VERSION : 0.1
   VAR
      HEADER : Struct
         DB_NR : Int := 3701;
         MIN_NR_EMS : Int := 1;
         MAX_NR_EMS : Int := 200;
         START_EMS : Int := 20;
         LAENGE_EMS_FLAGS : Int := 2;
         ACT_COUNT : Int := 0;
         Res120 : Int := 0;
         Res140 : Int := 0;
         Res160 : Int := 0;
         Res180 : Int := 0;
      END_STRUCT;
      EMS : Array[1..200] of "UDT_SDC_EMS_FLAGS";
      LADDR_EMS : Array[1..200] of HW_ANY;
   END_VAR
BEGIN
   EMS[3].SIMULATION := FALSE;
   EMS[2].SIMULATION := FALSE;
   EMS[200].FAULTY := TRUE;
   EMS[199].FAULTY := TRUE;
   EMS[198].FAULTY := TRUE;
   EMS[197].FAULTY := TRUE;
   EMS[196].FAULTY := TRUE;
   EMS[195].FAULTY := TRUE;
   EMS[194].FAULTY := TRUE;
   EMS[193].FAULTY := TRUE;
   EMS[192].FAULTY := TRUE;
   EMS[191].FAULTY := TRUE;
   EMS[190].FAULTY := TRUE;
   EMS[189].FAULTY := TRUE;
   EMS[188].FAULTY := TRUE;
   EMS[187].FAULTY := TRUE;
   EMS[186].FAULTY := TRUE;
   EMS[185].FAULTY := TRUE;
   EMS[184].FAULTY := TRUE;
   EMS[183].FAULTY := TRUE;
   EMS[182].FAULTY := TRUE;
   EMS[181].FAULTY := TRUE;
   EMS[180].FAULTY := TRUE;
   EMS[179].FAULTY := TRUE;
   EMS[178].FAULTY := TRUE;
   EMS[177].FAULTY := TRUE;
   EMS[176].FAULTY := TRUE;
   EMS[175].FAULTY := TRUE;
   EMS[174].FAULTY := TRUE;
   EMS[173].FAULTY := TRUE;
   EMS[172].FAULTY := TRUE;
   EMS[171].FAULTY := TRUE;
   EMS[170].FAULTY := TRUE;
   EMS[169].FAULTY := TRUE;
   EMS[168].FAULTY := TRUE;
   EMS[167].FAULTY := TRUE;
   EMS[166].FAULTY := TRUE;
   EMS[165].FAULTY := TRUE;
   EMS[164].FAULTY := TRUE;
   EMS[163].FAULTY := TRUE;
   EMS[162].FAULTY := TRUE;
   EMS[161].FAULTY := TRUE;
   EMS[160].FAULTY := TRUE;
   EMS[159].FAULTY := TRUE;
   EMS[158].FAULTY := TRUE;
   EMS[157].FAULTY := TRUE;
   EMS[156].FAULTY := TRUE;
   EMS[155].FAULTY := TRUE;
   EMS[154].FAULTY := TRUE;
   EMS[153].FAULTY := TRUE;
   EMS[152].FAULTY := TRUE;
   EMS[151].FAULTY := TRUE;
   EMS[150].FAULTY := TRUE;
   EMS[149].FAULTY := TRUE;
   EMS[148].FAULTY := TRUE;
   EMS[147].FAULTY := TRUE;
   EMS[146].FAULTY := TRUE;
   EMS[145].FAULTY := TRUE;
   EMS[144].FAULTY := TRUE;
   EMS[143].FAULTY := TRUE;
   EMS[142].FAULTY := TRUE;
   EMS[141].FAULTY := TRUE;
   EMS[140].FAULTY := TRUE;
   EMS[139].FAULTY := TRUE;
   EMS[138].FAULTY := TRUE;
   EMS[137].FAULTY := TRUE;
   EMS[136].FAULTY := TRUE;
   EMS[135].FAULTY := TRUE;
   EMS[134].FAULTY := TRUE;
   EMS[133].FAULTY := TRUE;
   EMS[132].FAULTY := TRUE;
   EMS[131].FAULTY := TRUE;
   EMS[130].FAULTY := TRUE;
   EMS[129].FAULTY := TRUE;
   EMS[128].FAULTY := TRUE;
   EMS[127].FAULTY := TRUE;
   EMS[126].FAULTY := TRUE;
   EMS[125].FAULTY := TRUE;
   EMS[124].FAULTY := TRUE;
   EMS[123].FAULTY := TRUE;
   EMS[122].FAULTY := TRUE;
   EMS[121].FAULTY := TRUE;
   EMS[120].FAULTY := TRUE;
   EMS[119].FAULTY := TRUE;
   EMS[118].FAULTY := TRUE;
   EMS[117].FAULTY := TRUE;
   EMS[116].FAULTY := TRUE;
   EMS[115].FAULTY := TRUE;
   EMS[114].FAULTY := TRUE;
   EMS[113].FAULTY := TRUE;
   EMS[112].FAULTY := TRUE;
   EMS[111].FAULTY := TRUE;
   EMS[110].FAULTY := TRUE;
   EMS[109].FAULTY := TRUE;
   EMS[108].FAULTY := TRUE;
   EMS[107].FAULTY := TRUE;
   EMS[106].FAULTY := TRUE;
   EMS[105].FAULTY := TRUE;
   EMS[104].FAULTY := TRUE;
   EMS[103].FAULTY := TRUE;
   EMS[102].FAULTY := TRUE;
   EMS[101].FAULTY := TRUE;
   EMS[100].FAULTY := TRUE;
   EMS[99].FAULTY := TRUE;
   EMS[98].FAULTY := TRUE;
   EMS[97].FAULTY := TRUE;
   EMS[96].FAULTY := TRUE;
   EMS[95].FAULTY := TRUE;
   EMS[94].FAULTY := TRUE;
   EMS[93].FAULTY := TRUE;
   EMS[92].FAULTY := TRUE;
   EMS[91].FAULTY := TRUE;
   EMS[90].FAULTY := TRUE;
   EMS[89].FAULTY := TRUE;
   EMS[88].FAULTY := TRUE;
   EMS[87].FAULTY := TRUE;
   EMS[86].FAULTY := TRUE;
   EMS[85].FAULTY := TRUE;
   EMS[84].FAULTY := TRUE;
   EMS[83].FAULTY := TRUE;
   EMS[82].FAULTY := TRUE;
   EMS[81].FAULTY := TRUE;
   EMS[80].FAULTY := TRUE;
   EMS[79].FAULTY := TRUE;
   EMS[78].FAULTY := TRUE;
   EMS[77].FAULTY := TRUE;
   EMS[76].FAULTY := TRUE;
   EMS[75].FAULTY := TRUE;
   EMS[74].FAULTY := TRUE;
   EMS[73].FAULTY := TRUE;
   EMS[72].FAULTY := TRUE;
   EMS[71].FAULTY := TRUE;
   EMS[70].FAULTY := TRUE;
   EMS[69].FAULTY := TRUE;
   EMS[68].FAULTY := TRUE;
   EMS[67].FAULTY := TRUE;
   EMS[66].FAULTY := TRUE;
   EMS[65].FAULTY := TRUE;
   EMS[64].FAULTY := TRUE;
   EMS[63].FAULTY := TRUE;
   EMS[62].FAULTY := TRUE;
   EMS[61].FAULTY := TRUE;
   EMS[60].FAULTY := TRUE;
   EMS[59].FAULTY := TRUE;
   EMS[58].FAULTY := TRUE;
   EMS[57].FAULTY := TRUE;
   EMS[56].FAULTY := TRUE;
   EMS[55].FAULTY := TRUE;
   EMS[54].FAULTY := FALSE;
   EMS[53].FAULTY := TRUE;
   EMS[52].FAULTY := TRUE;
   EMS[51].FAULTY := TRUE;
   EMS[50].FAULTY := TRUE;
   EMS[49].FAULTY := TRUE;
   EMS[48].FAULTY := TRUE;
   EMS[47].FAULTY := TRUE;
   EMS[46].FAULTY := TRUE;
   EMS[45].FAULTY := TRUE;
   EMS[44].FAULTY := TRUE;
   EMS[43].FAULTY := TRUE;
   EMS[42].FAULTY := TRUE;
   EMS[41].FAULTY := TRUE;
   EMS[40].FAULTY := TRUE;
   EMS[39].FAULTY := TRUE;
   EMS[38].FAULTY := TRUE;
   EMS[37].FAULTY := TRUE;
   EMS[36].FAULTY := TRUE;
   EMS[35].FAULTY := TRUE;
   EMS[34].FAULTY := FALSE;
   EMS[33].FAULTY := TRUE;
   EMS[32].FAULTY := FALSE;
   EMS[31].FAULTY := TRUE;
   EMS[30].FAULTY := TRUE;
   EMS[29].FAULTY := FALSE;
   EMS[28].FAULTY := TRUE;
   EMS[27].FAULTY := TRUE;
   EMS[26].FAULTY := TRUE;
   EMS[25].FAULTY := TRUE;
   EMS[24].FAULTY := TRUE;
   EMS[23].FAULTY := TRUE;
   EMS[22].FAULTY := TRUE;
   EMS[21].FAULTY := TRUE;
   EMS[20].FAULTY := TRUE;
   EMS[19].FAULTY := TRUE;
   EMS[18].FAULTY := TRUE;
   EMS[17].FAULTY := TRUE;
   EMS[16].FAULTY := TRUE;
   EMS[15].FAULTY := TRUE;
   EMS[14].FAULTY := TRUE;
   EMS[13].FAULTY := TRUE;
   EMS[12].FAULTY := TRUE;
   EMS[11].FAULTY := TRUE;
   EMS[10].FAULTY := TRUE;
   EMS[9].FAULTY := TRUE;
   EMS[8].FAULTY := TRUE;
   EMS[7].FAULTY := TRUE;
   EMS[6].FAULTY := TRUE;
   EMS[5].FAULTY := TRUE;
   EMS[4].FAULTY := TRUE;
   EMS[3].FAULTY := TRUE;
   // 3200 more start values not shown
END_DATA_BLOCK

DATA_BLOCK "DB_SDC_TS_PARAMETER_1"   // DB3704
{ S7_Optimized_Access := 'FALSE' }
AUTHOR : FFM
FAMILY : SDC
NAME : SECT_DEF
VERSION : 1.0
   VAR
      HEADER : Struct
         DB_NR : Int := 3704;
         MIN_NR_SEK : Int := 1;
         MAX_NR_SEK : Int := 100;
         START_DAT : Int := 20;
         LAENGE_SEK_DATA : Int := 260;
         ANZ_PROFIL : Int := 10;
         OFFEST_PROFIL : Int := 40;
         LAENGE_PROFIL_DATA : Int := 22;
         Res160 : Int := 0;
         Res : Int := 0;
      END_STRUCT;
      TS : Array[1..100] of "UDT_SDC_TS_PARAMETER";
   END_VAR
BEGIN
   TS[100].ALLG.Drive_speed_2 := 15000;
   TS[100].ALLG.Drive_speed_1 := 15000;
   TS[100].ALLG.Stop_Position := 2674;
   TS[100].ALLG.POS.End_1 := 371999;
   TS[100].ALLG.POS.Start_1 := 365500;
   TS[96].ALLG.Drive_speed_2 := 10000;
   TS[96].ALLG.Drive_speed_1 := 15000;
   TS[96].ALLG.Stop_Position := 3000;
   TS[96].ALLG.POS.End_1 := 365499;
   TS[96].ALLG.POS.Start_1 := 357900;
   TS[95].ALLG.Drive_speed_2 := 10000;
   TS[95].ALLG.Drive_speed_1 := 15000;
   TS[95].ALLG.Stop_Position := 3000;
   TS[95].ALLG.POS.End_1 := 357899;
   TS[95].ALLG.POS.Start_1 := 351800;
   TS[94].ALLG.Drive_speed_2 := 10000;
   TS[94].ALLG.Drive_speed_1 := 15000;
   TS[94].ALLG.Stop_Position := 3000;
   TS[94].ALLG.POS.End_1 := 351799;
   TS[94].ALLG.POS.Start_1 := 345700;
   TS[93].ALLG.Drive_speed_2 := 10000;
   TS[93].ALLG.Drive_speed_1 := 15000;
   TS[93].ALLG.Stop_Position := 3000;
   TS[93].ALLG.POS.End_1 := 345699;
   TS[93].ALLG.POS.Start_1 := 339600;
   TS[92].ALLG.Drive_speed_2 := 10000;
   TS[92].ALLG.Drive_speed_1 := 15000;
   TS[92].ALLG.Stop_Position := 3000;
   TS[92].ALLG.POS.End_1 := 339599;
   TS[92].ALLG.POS.Start_1 := 333500;
   TS[91].ALLG.Drive_speed_2 := 10000;
   TS[91].ALLG.Drive_speed_1 := 15000;
   TS[91].ALLG.Stop_Position := 3000;
   TS[91].ALLG.POS.End_1 := 333499;
   TS[91].ALLG.POS.Start_1 := 327400;
   TS[90].ALLG.Drive_speed_2 := 10000;
   TS[90].ALLG.Drive_speed_1 := 15000;
   TS[90].ALLG.Stop_Position := 3000;
   TS[90].ALLG.POS.End_1 := 327399;
   TS[90].ALLG.POS.Start_1 := 321300;
   TS[89].ALLG.Drive_speed_2 := 10000;
   TS[89].ALLG.Drive_speed_1 := 15000;
   TS[89].ALLG.Stop_Position := 3000;
   TS[89].ALLG.POS.End_1 := 321299;
   TS[89].ALLG.POS.Start_1 := 315200;
   TS[88].ALLG.Drive_speed_2 := 10000;
   TS[88].ALLG.Drive_speed_1 := 15000;
   TS[88].ALLG.Stop_Position := 3000;
   TS[88].ALLG.POS.End_1 := 315199;
   TS[88].ALLG.POS.Start_1 := 309100;
   TS[87].ALLG.Drive_speed_2 := 10000;
   TS[87].ALLG.Drive_speed_1 := 15000;
   TS[87].ALLG.Stop_Position := 3000;
   TS[87].ALLG.POS.End_1 := 309099;
   TS[87].ALLG.POS.Start_1 := 303000;
   TS[86].ALLG.Drive_speed_2 := 10000;
   TS[86].ALLG.Drive_speed_1 := 15000;
   TS[86].ALLG.POS.End_1 := 302999;
   TS[86].ALLG.POS.Start_1 := 300000;
   TS[1].ALLG.SEK_NEXT_1 := 0;
   TS[1].ALLG.SEK_NEXT_2 := 0;
   TS[1].ALLG.Spare[4] := 16#00;
   TS[1].ALLG.Spare[5] := 16#00;
   TS[1].ALLG.POS.Start_1 := 1687400;
   TS[1].ALLG.POS.End_1 := 1693799;
   TS[1].ALLG.POS.Start_2 := 0;
   TS[1].ALLG.POS.End_2 := 0;
   TS[1].ALLG.POS.Actionpoint_1 := 0;
   TS[1].ALLG.POS.Actionpoint_2 := 0;
   TS[1].ALLG.FLAGS.DIST_VAL[0] := FALSE;
   TS[1].ALLG.FLAGS.DIST_VAL[1] := FALSE;
   TS[1].ALLG.FLAGS.DIST_VAL[2] := FALSE;
   TS[1].ALLG.FLAGS.DIST_VAL[3] := FALSE;
   TS[1].ALLG.FLAGS.DIST_VAL[4] := FALSE;
   TS[1].ALLG.FLAGS.DIST_VAL[5] := FALSE;
   TS[1].ALLG.FLAGS.DIST_VAL[6] := FALSE;
   TS[1].ALLG.FLAGS.DIST_VAL[7] := FALSE;
   TS[1].ALLG.FLAGS.DIST_VAL[8] := FALSE;
   TS[1].ALLG.FLAGS.DIST_VAL[9] := TRUE;
   TS[1].ALLG.FLAGS.DIST_VAL[10] := FALSE;
   TS[1].ALLG.FLAGS.DIST_VAL[11] := FALSE;
   TS[1].ALLG.FLAGS.DIST_VAL[12] := FALSE;
   TS[1].ALLG.FLAGS.DIST_VAL[13] := FALSE;
   TS[1].ALLG.FLAGS.DIST_VAL[14] := FALSE;
   TS[1].ALLG.FLAGS.DIST_VAL[15] := FALSE;
   TS[1].ALLG.FLAGS.one_profile := FALSE;
   TS[1].ALLG.FLAGS.BLIND := FALSE;
   TS[1].ALLG.FLAGS.NO_DIST_CONT := FALSE;
   TS[1].ALLG.FLAGS.SYNCH_AREA := FALSE;
   TS[1].ALLG.FLAGS.bit24 := FALSE;
   TS[1].ALLG.FLAGS.bit25 := FALSE;
   TS[1].ALLG.FLAGS.bit26 := FALSE;
   TS[1].ALLG.FLAGS.bit27 := FALSE;
   TS[1].ALLG.FLAGS.EN_HOIST := FALSE;
   TS[1].ALLG.FLAGS.D_RESET_AFTER := FALSE;
   TS[1].ALLG.FLAGS.D_PULK := FALSE;
   TS[1].ALLG.FLAGS.bit33 := FALSE;
   TS[1].ALLG.FLAGS.bit34 := FALSE;
   TS[1].ALLG.FLAGS.bit35 := FALSE;
   TS[1].ALLG.FLAGS.bit36 := FALSE;
   TS[1].ALLG.FLAGS.Deutronic_ON := FALSE;
   TS[1].ALLG.Stop_Position := 5800;
   TS[1].ALLG.Drive_speed_1 := 15000;
   TS[1].ALLG.Drive_speed_2 := 6000;
   TS[1].PROFIL[1].Hoist_Pos_start := 0;
   TS[1].PROFIL[1].Height := 3890;
   TS[1].PROFIL[1].Hoist_speed := 2000;
   TS[1].PROFIL[1].Hoist_offset_1 := 0;
   TS[1].PROFIL[1].Hoist_offset_2 := 0;
   TS[1].PROFIL[1].Hoist_offset_3 := 0;
   TS[1].PROFIL[1].Hoist_offset_4 := 0;
   TS[1].PROFIL[1].Hoist_Start_offset_1 := 0;
   TS[1].PROFIL[1].Hoist_Start_offset_2 := 0;
   TS[1].PROFIL[1].Hoist_Start_offset_3 := 0;
   TS[1].PROFIL[1].Hoist_Start_offset_4 := 0;
   TS[1].PROFIL[2].Hoist_Pos_start := 0;
   TS[1].PROFIL[2].Height := 3890;
   TS[1].PROFIL[2].Hoist_speed := 2000;
   TS[1].PROFIL[2].Hoist_offset_1 := 0;
   TS[1].PROFIL[2].Hoist_offset_2 := 0;
   TS[1].PROFIL[2].Hoist_offset_3 := 0;
   TS[1].PROFIL[2].Hoist_offset_4 := 0;
   TS[1].PROFIL[2].Hoist_Start_offset_1 := 0;
   TS[1].PROFIL[2].Hoist_Start_offset_2 := 0;
   TS[1].PROFIL[2].Hoist_Start_offset_3 := 0;
   TS[1].PROFIL[2].Hoist_Start_offset_4 := 0;
   TS[1].PROFIL[3].Hoist_Pos_start := 0;
   TS[1].PROFIL[3].Height := 3890;
   TS[1].PROFIL[3].Hoist_speed := 2000;
   TS[1].PROFIL[3].Hoist_offset_1 := 0;
   TS[1].PROFIL[3].Hoist_offset_2 := 0;
   TS[1].PROFIL[3].Hoist_offset_3 := 0;
   TS[1].PROFIL[3].Hoist_offset_4 := 0;
   TS[1].PROFIL[3].Hoist_Start_offset_1 := 0;
   TS[1].PROFIL[3].Hoist_Start_offset_2 := 0;
   TS[1].PROFIL[3].Hoist_Start_offset_3 := 0;
   TS[1].PROFIL[3].Hoist_Start_offset_4 := 0;
   TS[1].PROFIL[4].Hoist_Pos_start := 0;
   TS[1].PROFIL[4].Height := 3890;
   TS[1].PROFIL[4].Hoist_speed := 2000;
   TS[1].PROFIL[4].Hoist_offset_1 := 0;
   TS[1].PROFIL[4].Hoist_offset_2 := 0;
   TS[1].PROFIL[4].Hoist_offset_3 := 0;
   TS[1].PROFIL[4].Hoist_offset_4 := 0;
   TS[1].PROFIL[4].Hoist_Start_offset_1 := 0;
   TS[1].PROFIL[4].Hoist_Start_offset_2 := 0;
   TS[1].PROFIL[4].Hoist_Start_offset_3 := 0;
   TS[1].PROFIL[4].Hoist_Start_offset_4 := 0;
   TS[1].PROFIL[5].Hoist_Pos_start := 0;
   TS[1].PROFIL[5].Height := 3890;
   TS[1].PROFIL[5].Hoist_speed := 2000;
   TS[1].PROFIL[5].Hoist_offset_1 := 0;
   TS[1].PROFIL[5].Hoist_offset_2 := 0;
   TS[1].PROFIL[5].Hoist_offset_3 := 0;
   TS[1].PROFIL[5].Hoist_offset_4 := 0;
   TS[1].PROFIL[5].Hoist_Start_offset_1 := 0;
   TS[1].PROFIL[5].Hoist_Start_offset_2 := 0;
   TS[1].PROFIL[5].Hoist_Start_offset_3 := 0;
   TS[1].PROFIL[5].Hoist_Start_offset_4 := 0;
   TS[1].PROFIL[6].Hoist_Pos_start := 0;
   TS[1].PROFIL[6].Height := 3890;
   TS[1].PROFIL[6].Hoist_speed := 2000;
   TS[1].PROFIL[6].Hoist_offset_1 := 0;
   TS[1].PROFIL[6].Hoist_offset_2 := 0;
   TS[1].PROFIL[6].Hoist_offset_3 := 0;
   TS[1].PROFIL[6].Hoist_offset_4 := 0;
   TS[1].PROFIL[6].Hoist_Start_offset_1 := 0;
   TS[1].PROFIL[6].Hoist_Start_offset_2 := 0;
   TS[1].PROFIL[6].Hoist_Start_offset_3 := 0;
   TS[1].PROFIL[6].Hoist_Start_offset_4 := 0;
   TS[1].PROFIL[7].Hoist_Pos_start := 0;
   TS[1].PROFIL[7].Height := 3890;
   TS[1].PROFIL[7].Hoist_speed := 2000;
   TS[1].PROFIL[7].Hoist_offset_1 := 0;
   TS[1].PROFIL[7].Hoist_offset_2 := 0;
   TS[1].PROFIL[7].Hoist_offset_3 := 0;
   TS[1].PROFIL[7].Hoist_offset_4 := 0;
   TS[1].PROFIL[7].Hoist_Start_offset_1 := 0;
   TS[1].PROFIL[7].Hoist_Start_offset_2 := 0;
   TS[1].PROFIL[7].Hoist_Start_offset_3 := 0;
   TS[1].PROFIL[7].Hoist_Start_offset_4 := 0;
   TS[1].PROFIL[8].Hoist_Pos_start := 0;
   TS[1].PROFIL[8].Height := 3890;
   TS[1].PROFIL[8].Hoist_speed := 2000;
   TS[1].PROFIL[8].Hoist_offset_1 := 0;
   TS[1].PROFIL[8].Hoist_offset_2 := 0;
   TS[1].PROFIL[8].Hoist_offset_3 := 0;
   TS[1].PROFIL[8].Hoist_offset_4 := 0;
   TS[1].PROFIL[8].Hoist_Start_offset_1 := 0;
   TS[1].PROFIL[8].Hoist_Start_offset_2 := 0;
   TS[1].PROFIL[8].Hoist_Start_offset_3 := 0;
   TS[1].PROFIL[8].Hoist_Start_offset_4 := 0;
   TS[1].PROFIL[9].Hoist_Pos_start := 0;
   TS[1].PROFIL[9].Height := 3890;
   TS[1].PROFIL[9].Hoist_speed := 2000;
   TS[1].PROFIL[9].Hoist_offset_1 := 0;
   TS[1].PROFIL[9].Hoist_offset_2 := 0;
   TS[1].PROFIL[9].Hoist_offset_3 := 0;
   TS[1].PROFIL[9].Hoist_offset_4 := 0;
   TS[1].PROFIL[9].Hoist_Start_offset_1 := 0;
   // 15300 more start values not shown
END_DATA_BLOCK

DATA_BLOCK "DB_SDC_TS_PARAMETER_2"   // DB3705
{ S7_Optimized_Access := 'FALSE' }
AUTHOR : FFM
FAMILY : SDC
NAME : SECT_DEF
VERSION : 1.0
   VAR
      HEADER : Struct
         DB_NR : Int := 3705;
         MIN_NR_SEK : Int := 101;
         MAX_NR_SEK : Int := 200;
         START_DAT : Int := 20;
         LAENGE_SEK_DATA : Int := 260;
         ANZ_PROFIL : Int := 10;
         OFFEST_PROFIL : Int := 40;
         LAENGE_PROFIL_DATA : Int := 22;
         Res160 : Int := 0;
         Res : Int := 0;
      END_STRUCT;
      TS : Array[101..200] of "UDT_SDC_TS_PARAMETER";
   END_VAR
BEGIN
   TS[101].ALLG.POS.Start_1 := 372000;
   TS[101].ALLG.POS.End_1 := 378499;
   TS[101].ALLG.Stop_Position := 3000;
   TS[101].ALLG.Drive_speed_1 := 20000;
   TS[101].ALLG.Drive_speed_2 := 20000;
   TS[102].ALLG.POS.Start_1 := 378500;
   TS[102].ALLG.POS.End_1 := 384999;
   TS[102].ALLG.Stop_Position := 3000;
   TS[102].ALLG.Drive_speed_1 := 10000;
   TS[102].ALLG.Drive_speed_2 := 7000;
   TS[103].ALLG.POS.Start_1 := 385000;
   TS[103].ALLG.POS.End_1 := 391499;
   TS[103].ALLG.Stop_Position := 3000;
   TS[103].ALLG.Drive_speed_1 := 20000;
   TS[103].ALLG.Drive_speed_2 := 20000;
   TS[104].ALLG.POS.Start_1 := 391500;
   TS[104].ALLG.POS.End_1 := 397999;
   TS[104].ALLG.Stop_Position := 3000;
   TS[104].ALLG.Drive_speed_1 := 20000;
   TS[104].ALLG.Drive_speed_2 := 20000;
   TS[105].ALLG.POS.Start_1 := 398000;
   TS[105].ALLG.POS.End_1 := 404499;
   TS[105].ALLG.Stop_Position := 3000;
   TS[105].ALLG.Drive_speed_1 := 22000;
   TS[105].ALLG.Drive_speed_2 := 20000;
   TS[106].ALLG.POS.Start_1 := 404500;
   TS[106].ALLG.POS.End_1 := 410999;
   TS[106].ALLG.Stop_Position := 3000;
   TS[106].ALLG.Drive_speed_1 := 22000;
   TS[106].ALLG.Drive_speed_2 := 5000;
   TS[107].ALLG.POS.Start_1 := 411000;
   TS[107].ALLG.POS.End_1 := 417499;
   TS[107].ALLG.Stop_Position := 3000;
   TS[107].ALLG.Drive_speed_1 := 18000;
   TS[107].ALLG.Drive_speed_2 := 4000;
   TS[108].ALLG.POS.Start_1 := 417500;
   TS[108].ALLG.POS.End_1 := 423999;
   TS[108].ALLG.Stop_Position := 3000;
   TS[108].ALLG.Drive_speed_1 := 22000;
   TS[108].ALLG.Drive_speed_2 := 10000;
   TS[109].ALLG.POS.Start_1 := 424000;
   TS[109].ALLG.POS.End_1 := 430499;
   TS[109].ALLG.Stop_Position := 3000;
   TS[109].ALLG.Drive_speed_1 := 20000;
   TS[109].ALLG.Drive_speed_2 := 10000;
   TS[110].ALLG.POS.Start_1 := 430500;
   TS[110].ALLG.POS.End_1 := 436999;
   TS[110].ALLG.Stop_Position := 2674;
   TS[110].ALLG.Drive_speed_1 := 15000;
   TS[110].ALLG.Drive_speed_2 := 10000;
   TS[111].ALLG.POS.Start_1 := 437000;
   TS[111].ALLG.POS.End_1 := 443499;
   TS[111].ALLG.Stop_Position := 3000;
   TS[111].ALLG.Drive_speed_1 := 15000;
   TS[111].ALLG.Drive_speed_2 := 10000;
   TS[120].ALLG.POS.Start_1 := 443500;
   TS[120].ALLG.POS.End_1 := 450499;
   TS[120].ALLG.Stop_Position := 5200;
   TS[120].ALLG.Drive_speed_1 := 15000;
   TS[120].ALLG.Drive_speed_2 := 10000;
   TS[121].ALLG.POS.Start_1 := 450500;
   TS[121].ALLG.POS.End_1 := 457499;
   TS[121].ALLG.Stop_Position := 5500;
   TS[121].ALLG.Drive_speed_1 := 15000;
   TS[121].ALLG.Drive_speed_2 := 10000;
   TS[122].ALLG.POS.Start_1 := 457500;
   TS[122].ALLG.POS.End_1 := 463999;
   TS[122].ALLG.Stop_Position := 5000;
   TS[122].ALLG.Drive_speed_1 := 15000;
   TS[122].ALLG.Drive_speed_2 := 10000;
   TS[123].ALLG.POS.Start_1 := 464000;
   TS[123].ALLG.POS.End_1 := 470499;
   TS[123].ALLG.Stop_Position := 5100;
   TS[123].ALLG.Drive_speed_1 := 15000;
   TS[123].ALLG.Drive_speed_2 := 10000;
   TS[124].ALLG.POS.Start_1 := 470500;
   TS[124].ALLG.POS.End_1 := 476999;
   TS[124].ALLG.Stop_Position := 5000;
   TS[124].ALLG.Drive_speed_1 := 15000;
   TS[124].ALLG.Drive_speed_2 := 10000;
   TS[125].ALLG.POS.Start_1 := 477000;
   TS[125].ALLG.POS.End_1 := 483999;
   TS[125].ALLG.Stop_Position := 6400;
   TS[125].ALLG.Drive_speed_1 := 15000;
   TS[125].ALLG.Drive_speed_2 := 10000;
   TS[126].ALLG.POS.Start_1 := 484000;
   TS[126].ALLG.POS.End_1 := 491999;
   TS[126].ALLG.Stop_Position := 7200;
   TS[126].ALLG.Drive_speed_1 := 15000;
   TS[126].ALLG.Drive_speed_2 := 10000;
   TS[127].ALLG.POS.Start_1 := 492000;
   TS[127].ALLG.POS.End_1 := 498199;
   TS[127].ALLG.Stop_Position := 5400;
   TS[127].ALLG.Drive_speed_1 := 15000;
   TS[127].ALLG.Drive_speed_2 := 10000;
   TS[128].ALLG.POS.Start_1 := 498200;
   TS[128].ALLG.POS.End_1 := 504399;
   TS[128].ALLG.Stop_Position := 2954;
   TS[128].ALLG.Drive_speed_1 := 15000;
   TS[128].ALLG.Drive_speed_2 := 10000;
   TS[129].ALLG.POS.Start_1 := 504400;
   TS[129].ALLG.POS.End_1 := 511399;
   TS[129].ALLG.Stop_Position := 6300;
   TS[129].ALLG.Drive_speed_1 := 15000;
   TS[129].ALLG.Drive_speed_2 := 10000;
   TS[130].ALLG.POS.Start_1 := 511400;
   TS[130].ALLG.POS.End_1 := 518399;
   TS[130].ALLG.Stop_Position := 6300;
   TS[130].ALLG.Drive_speed_1 := 15000;
   TS[130].ALLG.Drive_speed_2 := 10000;
   TS[131].ALLG.POS.Start_1 := 518400;
   TS[131].ALLG.POS.End_1 := 525599;
   TS[131].ALLG.Stop_Position := 6300;
   TS[131].ALLG.Drive_speed_1 := 15000;
   TS[131].ALLG.Drive_speed_2 := 10000;
   TS[132].ALLG.POS.Start_1 := 525600;
   TS[132].ALLG.POS.End_1 := 529699;
   TS[132].ALLG.Stop_Position := 4299;
   TS[132].ALLG.Drive_speed_1 := 10000;
   TS[132].ALLG.Drive_speed_2 := 10000;
   TS[140].ALLG.POS.Start_1 := 529700;
   TS[140].ALLG.POS.End_1 := 535699;
   TS[140].ALLG.Stop_Position := 5900;
   TS[140].ALLG.Drive_speed_1 := 30000;
   TS[140].ALLG.Drive_speed_2 := 10000;
   TS[141].ALLG.POS.Start_1 := 535700;
   TS[141].ALLG.POS.End_1 := 541699;
   TS[141].ALLG.Stop_Position := 5900;
   TS[141].ALLG.Drive_speed_1 := 30000;
   TS[141].ALLG.Drive_speed_2 := 10000;
   TS[142].ALLG.POS.Start_1 := 541700;
   TS[142].ALLG.POS.End_1 := 547699;
   TS[142].ALLG.Stop_Position := 5900;
   TS[142].ALLG.Drive_speed_1 := 30000;
   TS[142].ALLG.Drive_speed_2 := 10000;
   TS[143].ALLG.POS.Start_1 := 547700;
   TS[143].ALLG.POS.End_1 := 553699;
   TS[143].ALLG.Stop_Position := 5900;
   TS[143].ALLG.Drive_speed_1 := 30000;
   TS[143].ALLG.Drive_speed_2 := 10000;
   TS[144].ALLG.POS.Start_1 := 553700;
   TS[144].ALLG.POS.End_1 := 559699;
   TS[144].ALLG.Stop_Position := 5900;
   TS[144].ALLG.Drive_speed_1 := 30000;
   TS[144].ALLG.Drive_speed_2 := 10000;
   TS[145].ALLG.POS.Start_1 := 559700;
   TS[145].ALLG.POS.End_1 := 565699;
   TS[145].ALLG.Stop_Position := 5900;
   TS[145].ALLG.Drive_speed_1 := 30000;
   TS[145].ALLG.Drive_speed_2 := 10000;
   TS[146].ALLG.POS.Start_1 := 565700;
   TS[146].ALLG.POS.End_1 := 571699;
   TS[146].ALLG.Stop_Position := 5900;
   TS[146].ALLG.Drive_speed_1 := 30000;
   TS[146].ALLG.Drive_speed_2 := 10000;
   TS[147].ALLG.POS.Start_1 := 571700;
   TS[147].ALLG.POS.End_1 := 577699;
   TS[147].ALLG.Stop_Position := 5900;
   TS[147].ALLG.Drive_speed_1 := 30000;
   TS[147].ALLG.Drive_speed_2 := 10000;
   TS[148].ALLG.POS.Start_1 := 577700;
   TS[148].ALLG.POS.End_1 := 583699;
   TS[148].ALLG.Stop_Position := 5900;
   TS[148].ALLG.Drive_speed_1 := 30000;
   TS[148].ALLG.Drive_speed_2 := 10000;
   TS[149].ALLG.POS.Start_1 := 583700;
   TS[149].ALLG.POS.End_1 := 589699;
   TS[149].ALLG.Stop_Position := 5900;
   TS[149].ALLG.Drive_speed_1 := 30000;
   TS[149].ALLG.Drive_speed_2 := 10000;
   TS[150].ALLG.POS.Start_1 := 589700;
   TS[150].ALLG.POS.End_1 := 595699;
   TS[150].ALLG.Stop_Position := 5900;
   TS[150].ALLG.Drive_speed_1 := 25000;
   TS[150].ALLG.Drive_speed_2 := 10000;
   TS[151].ALLG.POS.Start_1 := 595700;
   TS[151].ALLG.POS.End_1 := 601699;
   TS[151].ALLG.Stop_Position := 5900;
   TS[151].ALLG.Drive_speed_1 := 18000;
   TS[151].ALLG.Drive_speed_2 := 10000;
   TS[152].ALLG.POS.Start_1 := 601700;
   TS[152].ALLG.POS.End_1 := 607699;
   TS[152].ALLG.Stop_Position := 5900;
   TS[152].ALLG.Drive_speed_1 := 18000;
   TS[152].ALLG.Drive_speed_2 := 10000;
   TS[160].ALLG.POS.Start_1 := 607700;
   TS[160].ALLG.POS.End_1 := 613699;
   TS[160].ALLG.Stop_Position := 5900;
   TS[160].ALLG.Drive_speed_1 := 20000;
   TS[160].ALLG.Drive_speed_2 := 10000;
   TS[161].ALLG.POS.Start_1 := 613700;
   TS[161].ALLG.POS.End_1 := 619699;
   TS[161].ALLG.Stop_Position := 5900;
   TS[161].ALLG.Drive_speed_1 := 20000;
   TS[161].ALLG.Drive_speed_2 := 10000;
   TS[162].ALLG.POS.Start_1 := 619700;
   TS[162].ALLG.POS.End_1 := 625699;
   TS[162].ALLG.Stop_Position := 5900;
   TS[162].ALLG.Drive_speed_1 := 20000;
   TS[162].ALLG.Drive_speed_2 := 10000;
   // 15300 more start values not shown
END_DATA_BLOCK

DATA_BLOCK "DB_SDC_TS_PARAMETER_3"   // DB3706
{ S7_Optimized_Access := 'FALSE' }
AUTHOR : FFM
FAMILY : SDC
NAME : SECT_DEF
VERSION : 1.0
   VAR
      HEADER : Struct   // Struktur für Datenheader // nicht verschieben
         DB_NR : Int := 3706;   // DB Nummer
         MIN_NR_SEK : Int := 201;   // Niedrigste SEK Nummer im DB
         MAX_NR_SEK : Int := 300;   // Höchste SEK Nummer im DB
         START_DAT : Int := 20;   // Startadresse der SEK im DB
         LAENGE_SEK_DATA : Int := 260;   // Länge SEK Data
         ANZ_PROFIL : Int := 10;   // Number of Profiles
         OFFEST_PROFIL : Int := 40;   // Offestadresse der Profilparameter im TS-Parameterdatensatz
         LAENGE_PROFIL_DATA : Int := 22;   // Länge SEK Data
         Res160 : Int := 0;   // Reserve
         Res : Int := 0;   // Reserve
      END_STRUCT;
      TS : Array[201..300] of "UDT_SDC_TS_PARAMETER";
   END_VAR
BEGIN
   TS[201].ALLG.SEK_NEXT_1 := 0;
   TS[201].ALLG.SEK_NEXT_2 := 0;
   TS[201].ALLG.Spare[4] := 16#00;
   TS[201].ALLG.Spare[5] := 16#00;
   TS[201].ALLG.POS.Start_1 := 709550;
   TS[201].ALLG.POS.End_1 := 715849;
   TS[201].ALLG.POS.Start_2 := 0;
   TS[201].ALLG.POS.End_2 := 0;
   TS[201].ALLG.POS.Actionpoint_1 := 0;
   TS[201].ALLG.POS.Actionpoint_2 := 0;
   TS[201].ALLG.FLAGS.DIST_VAL[0] := FALSE;
   TS[201].ALLG.FLAGS.DIST_VAL[1] := FALSE;
   TS[201].ALLG.FLAGS.DIST_VAL[2] := FALSE;
   TS[201].ALLG.FLAGS.DIST_VAL[3] := FALSE;
   TS[201].ALLG.FLAGS.DIST_VAL[4] := FALSE;
   TS[201].ALLG.FLAGS.DIST_VAL[5] := FALSE;
   TS[201].ALLG.FLAGS.DIST_VAL[6] := FALSE;
   TS[201].ALLG.FLAGS.DIST_VAL[7] := FALSE;
   TS[201].ALLG.FLAGS.DIST_VAL[8] := FALSE;
   TS[201].ALLG.FLAGS.DIST_VAL[9] := TRUE;
   TS[201].ALLG.FLAGS.DIST_VAL[10] := FALSE;
   TS[201].ALLG.FLAGS.DIST_VAL[11] := FALSE;
   TS[201].ALLG.FLAGS.DIST_VAL[12] := FALSE;
   TS[201].ALLG.FLAGS.DIST_VAL[13] := FALSE;
   TS[201].ALLG.FLAGS.DIST_VAL[14] := FALSE;
   TS[201].ALLG.FLAGS.DIST_VAL[15] := FALSE;
   TS[201].ALLG.FLAGS.one_profile := FALSE;
   TS[201].ALLG.FLAGS.BLIND := FALSE;
   TS[201].ALLG.FLAGS.NO_DIST_CONT := FALSE;
   TS[201].ALLG.FLAGS.SYNCH_AREA := FALSE;
   TS[201].ALLG.FLAGS.bit24 := FALSE;
   TS[201].ALLG.FLAGS.bit25 := FALSE;
   TS[201].ALLG.FLAGS.bit26 := FALSE;
   TS[201].ALLG.FLAGS.bit27 := FALSE;
   TS[201].ALLG.FLAGS.EN_HOIST := FALSE;
   TS[201].ALLG.FLAGS.D_RESET_AFTER := FALSE;
   TS[201].ALLG.FLAGS.D_PULK := FALSE;
   TS[201].ALLG.FLAGS.bit33 := FALSE;
   TS[201].ALLG.FLAGS.bit34 := FALSE;
   TS[201].ALLG.FLAGS.bit35 := FALSE;
   TS[201].ALLG.FLAGS.bit36 := FALSE;
   TS[201].ALLG.FLAGS.Deutronic_ON := FALSE;
   TS[201].ALLG.Stop_Position := 5800;
   TS[201].ALLG.Drive_speed_1 := 18000;
   TS[201].ALLG.Drive_speed_2 := 6000;
   TS[201].PROFIL[1].Hoist_Pos_start := 0;
   TS[201].PROFIL[1].Height := 3890;
   TS[201].PROFIL[1].Hoist_speed := 2000;
   TS[201].PROFIL[1].Hoist_offset_1 := 0;
   TS[201].PROFIL[1].Hoist_offset_2 := 0;
   TS[201].PROFIL[1].Hoist_offset_3 := 0;
   TS[201].PROFIL[1].Hoist_offset_4 := 0;
   TS[201].PROFIL[1].Hoist_Start_offset_1 := 0;
   TS[201].PROFIL[1].Hoist_Start_offset_2 := 0;
   TS[201].PROFIL[1].Hoist_Start_offset_3 := 0;
   TS[201].PROFIL[1].Hoist_Start_offset_4 := 0;
   TS[201].PROFIL[2].Hoist_Pos_start := 0;
   TS[201].PROFIL[2].Height := 3890;
   TS[201].PROFIL[2].Hoist_speed := 2000;
   TS[201].PROFIL[2].Hoist_offset_1 := 0;
   TS[201].PROFIL[2].Hoist_offset_2 := 0;
   TS[201].PROFIL[2].Hoist_offset_3 := 0;
   TS[201].PROFIL[2].Hoist_offset_4 := 0;
   TS[201].PROFIL[2].Hoist_Start_offset_1 := 0;
   TS[201].PROFIL[2].Hoist_Start_offset_2 := 0;
   TS[201].PROFIL[2].Hoist_Start_offset_3 := 0;
   TS[201].PROFIL[2].Hoist_Start_offset_4 := 0;
   TS[201].PROFIL[3].Hoist_Pos_start := 0;
   TS[201].PROFIL[3].Height := 3890;
   TS[201].PROFIL[3].Hoist_speed := 2000;
   TS[201].PROFIL[3].Hoist_offset_1 := 0;
   TS[201].PROFIL[3].Hoist_offset_2 := 0;
   TS[201].PROFIL[3].Hoist_offset_3 := 0;
   TS[201].PROFIL[3].Hoist_offset_4 := 0;
   TS[201].PROFIL[3].Hoist_Start_offset_1 := 0;
   TS[201].PROFIL[3].Hoist_Start_offset_2 := 0;
   TS[201].PROFIL[3].Hoist_Start_offset_3 := 0;
   TS[201].PROFIL[3].Hoist_Start_offset_4 := 0;
   TS[201].PROFIL[4].Hoist_Pos_start := 0;
   TS[201].PROFIL[4].Height := 3890;
   TS[201].PROFIL[4].Hoist_speed := 2000;
   TS[201].PROFIL[4].Hoist_offset_1 := 0;
   TS[201].PROFIL[4].Hoist_offset_2 := 0;
   TS[201].PROFIL[4].Hoist_offset_3 := 0;
   TS[201].PROFIL[4].Hoist_offset_4 := 0;
   TS[201].PROFIL[4].Hoist_Start_offset_1 := 0;
   TS[201].PROFIL[4].Hoist_Start_offset_2 := 0;
   TS[201].PROFIL[4].Hoist_Start_offset_3 := 0;
   TS[201].PROFIL[4].Hoist_Start_offset_4 := 0;
   TS[201].PROFIL[5].Hoist_Pos_start := 0;
   TS[201].PROFIL[5].Height := 3890;
   TS[201].PROFIL[5].Hoist_speed := 2000;
   TS[201].PROFIL[5].Hoist_offset_1 := 0;
   TS[201].PROFIL[5].Hoist_offset_2 := 0;
   TS[201].PROFIL[5].Hoist_offset_3 := 0;
   TS[201].PROFIL[5].Hoist_offset_4 := 0;
   TS[201].PROFIL[5].Hoist_Start_offset_1 := 0;
   TS[201].PROFIL[5].Hoist_Start_offset_2 := 0;
   TS[201].PROFIL[5].Hoist_Start_offset_3 := 0;
   TS[201].PROFIL[5].Hoist_Start_offset_4 := 0;
   TS[201].PROFIL[6].Hoist_Pos_start := 0;
   TS[201].PROFIL[6].Height := 3890;
   TS[201].PROFIL[6].Hoist_speed := 2000;
   TS[201].PROFIL[6].Hoist_offset_1 := 0;
   TS[201].PROFIL[6].Hoist_offset_2 := 0;
   TS[201].PROFIL[6].Hoist_offset_3 := 0;
   TS[201].PROFIL[6].Hoist_offset_4 := 0;
   TS[201].PROFIL[6].Hoist_Start_offset_1 := 0;
   TS[201].PROFIL[6].Hoist_Start_offset_2 := 0;
   TS[201].PROFIL[6].Hoist_Start_offset_3 := 0;
   TS[201].PROFIL[6].Hoist_Start_offset_4 := 0;
   TS[201].PROFIL[7].Hoist_Pos_start := 0;
   TS[201].PROFIL[7].Height := 3890;
   TS[201].PROFIL[7].Hoist_speed := 2000;
   TS[201].PROFIL[7].Hoist_offset_1 := 0;
   TS[201].PROFIL[7].Hoist_offset_2 := 0;
   TS[201].PROFIL[7].Hoist_offset_3 := 0;
   TS[201].PROFIL[7].Hoist_offset_4 := 0;
   TS[201].PROFIL[7].Hoist_Start_offset_1 := 0;
   TS[201].PROFIL[7].Hoist_Start_offset_2 := 0;
   TS[201].PROFIL[7].Hoist_Start_offset_3 := 0;
   TS[201].PROFIL[7].Hoist_Start_offset_4 := 0;
   TS[201].PROFIL[8].Hoist_Pos_start := 0;
   TS[201].PROFIL[8].Height := 3890;
   TS[201].PROFIL[8].Hoist_speed := 2000;
   TS[201].PROFIL[8].Hoist_offset_1 := 0;
   TS[201].PROFIL[8].Hoist_offset_2 := 0;
   TS[201].PROFIL[8].Hoist_offset_3 := 0;
   TS[201].PROFIL[8].Hoist_offset_4 := 0;
   TS[201].PROFIL[8].Hoist_Start_offset_1 := 0;
   TS[201].PROFIL[8].Hoist_Start_offset_2 := 0;
   TS[201].PROFIL[8].Hoist_Start_offset_3 := 0;
   TS[201].PROFIL[8].Hoist_Start_offset_4 := 0;
   TS[201].PROFIL[9].Hoist_Pos_start := 0;
   TS[201].PROFIL[9].Height := 3890;
   TS[201].PROFIL[9].Hoist_speed := 2000;
   TS[201].PROFIL[9].Hoist_offset_1 := 0;
   TS[201].PROFIL[9].Hoist_offset_2 := 0;
   TS[201].PROFIL[9].Hoist_offset_3 := 0;
   TS[201].PROFIL[9].Hoist_offset_4 := 0;
   TS[201].PROFIL[9].Hoist_Start_offset_1 := 0;
   TS[201].PROFIL[9].Hoist_Start_offset_2 := 0;
   TS[201].PROFIL[9].Hoist_Start_offset_3 := 0;
   TS[201].PROFIL[9].Hoist_Start_offset_4 := 0;
   TS[201].PROFIL[10].Hoist_Pos_start := 0;
   TS[201].PROFIL[10].Height := 3890;
   TS[201].PROFIL[10].Hoist_speed := 2000;
   TS[201].PROFIL[10].Hoist_offset_1 := 0;
   TS[201].PROFIL[10].Hoist_offset_2 := 0;
   TS[201].PROFIL[10].Hoist_offset_3 := 0;
   TS[201].PROFIL[10].Hoist_offset_4 := 0;
   TS[201].PROFIL[10].Hoist_Start_offset_1 := 0;
   TS[201].PROFIL[10].Hoist_Start_offset_2 := 0;
   TS[201].PROFIL[10].Hoist_Start_offset_3 := 0;
   TS[201].PROFIL[10].Hoist_Start_offset_4 := 0;
   TS[202].ALLG.SEK_NEXT_1 := 0;
   TS[202].ALLG.SEK_NEXT_2 := 0;
   TS[202].ALLG.Spare[4] := 16#00;
   TS[202].ALLG.Spare[5] := 16#00;
   TS[202].ALLG.POS.Start_1 := 715850;
   TS[202].ALLG.POS.End_1 := 722149;
   TS[202].ALLG.POS.Start_2 := 0;
   TS[202].ALLG.POS.End_2 := 0;
   TS[202].ALLG.POS.Actionpoint_1 := 0;
   TS[202].ALLG.POS.Actionpoint_2 := 0;
   TS[202].ALLG.FLAGS.DIST_VAL[0] := FALSE;
   TS[202].ALLG.FLAGS.DIST_VAL[1] := FALSE;
   TS[202].ALLG.FLAGS.DIST_VAL[2] := FALSE;
   TS[202].ALLG.FLAGS.DIST_VAL[3] := FALSE;
   TS[202].ALLG.FLAGS.DIST_VAL[4] := FALSE;
   TS[202].ALLG.FLAGS.DIST_VAL[5] := FALSE;
   TS[202].ALLG.FLAGS.DIST_VAL[6] := FALSE;
   TS[202].ALLG.FLAGS.DIST_VAL[7] := FALSE;
   TS[202].ALLG.FLAGS.DIST_VAL[8] := FALSE;
   TS[202].ALLG.FLAGS.DIST_VAL[9] := TRUE;
   TS[202].ALLG.FLAGS.DIST_VAL[10] := FALSE;
   TS[202].ALLG.FLAGS.DIST_VAL[11] := FALSE;
   TS[202].ALLG.FLAGS.DIST_VAL[12] := FALSE;
   TS[202].ALLG.FLAGS.DIST_VAL[13] := FALSE;
   TS[202].ALLG.FLAGS.DIST_VAL[14] := FALSE;
   TS[202].ALLG.FLAGS.DIST_VAL[15] := FALSE;
   TS[202].ALLG.FLAGS.one_profile := FALSE;
   TS[202].ALLG.FLAGS.BLIND := FALSE;
   TS[202].ALLG.FLAGS.NO_DIST_CONT := FALSE;
   TS[202].ALLG.FLAGS.SYNCH_AREA := FALSE;
   TS[202].ALLG.FLAGS.bit24 := FALSE;
   TS[202].ALLG.FLAGS.bit25 := FALSE;
   TS[202].ALLG.FLAGS.bit26 := FALSE;
   TS[202].ALLG.FLAGS.bit27 := FALSE;
   TS[202].ALLG.FLAGS.EN_HOIST := FALSE;
   TS[202].ALLG.FLAGS.D_RESET_AFTER := FALSE;
   TS[202].ALLG.FLAGS.D_PULK := FALSE;
   TS[202].ALLG.FLAGS.bit33 := FALSE;
   TS[202].ALLG.FLAGS.bit34 := FALSE;
   TS[202].ALLG.FLAGS.bit35 := FALSE;
   TS[202].ALLG.FLAGS.bit36 := FALSE;
   TS[202].ALLG.FLAGS.Deutronic_ON := FALSE;
   TS[202].ALLG.Stop_Position := 5800;
   TS[202].ALLG.Drive_speed_1 := 18000;
   TS[202].ALLG.Drive_speed_2 := 6000;
   // 15300 more start values not shown
END_DATA_BLOCK

